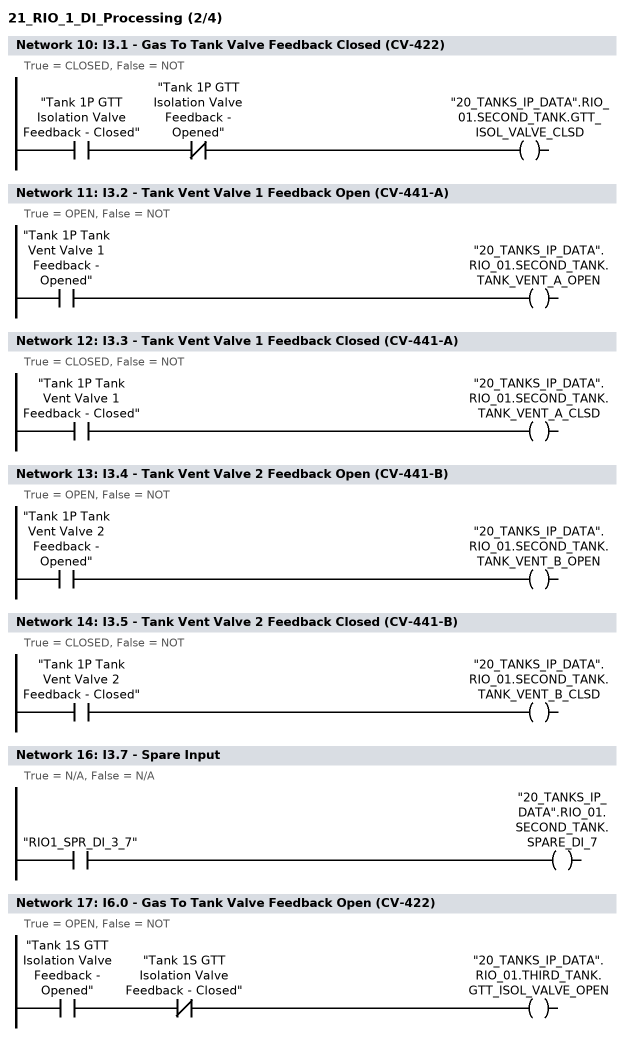
   RUNG wire#powerrail
      Contact( "Tank 1P GTT Isolation Valve Feedback - Closed" )
      I_Contact( "Tank 1P GTT Isolation Valve Feedback - Opened" )
      Coil( "20_TANKS_IP_DATA".RIO_01.SECOND_TANK.GTT_ISOL_VALVE_CLSD )
   END_RUNG
   // the same network as SCL:
   "20_TANKS_IP_DATA".RIO_01.SECOND_TANK.GTT_ISOL_VALVE_CLSD := "Tank 1P GTT Isolation Valve Feedback - Closed" AND NOT "Tank 1P GTT Isolation Valve Feedback - Opened";
END_REGION

REGION Network 11: I3.2 - Tank Vent Valve 1 Feedback Open (CV-441-A)
   // True = OPEN, False = NOT
   RUNG wire#powerrail
      Contact( "Tank 1P Tank Vent Valve 1 Feedback - Opened" )
      Coil( "20_TANKS_IP_DATA".RIO_01.SECOND_TANK.TANK_VENT_A_OPEN )
   END_RUNG
   // the same network as SCL:
   "20_TANKS_IP_DATA".RIO_01.SECOND_TANK.TANK_VENT_A_OPEN := "Tank 1P Tank Vent Valve 1 Feedback - Opened";
END_REGION

REGION Network 12: I3.3 - Tank Vent Valve 1 Feedback Closed (CV-441-A)
   // True = CLOSED, False = NOT
   RUNG wire#powerrail
      Contact( "Tank 1P Tank Vent Valve 1 Feedback - Closed" )
      Coil( "20_TANKS_IP_DATA".RIO_01.SECOND_TANK.TANK_VENT_A_CLSD )
   END_RUNG
   // the same network as SCL:
   "20_TANKS_IP_DATA".RIO_01.SECOND_TANK.TANK_VENT_A_CLSD := "Tank 1P Tank Vent Valve 1 Feedback - Closed";
END_REGION

REGION Network 13: I3.4 - Tank Vent Valve 2 Feedback Open (CV-441-B)
   // True = OPEN, False = NOT
   RUNG wire#powerrail
      Contact( "Tank 1P Tank Vent Valve 2 Feedback - Opened" )
      Coil( "20_TANKS_IP_DATA".RIO_01.SECOND_TANK.TANK_VENT_B_OPEN )
   END_RUNG
   // the same network as SCL:
   "20_TANKS_IP_DATA".RIO_01.SECOND_TANK.TANK_VENT_B_OPEN := "Tank 1P Tank Vent Valve 2 Feedback - Opened";
END_REGION

REGION Network 14: I3.5 - Tank Vent Valve 2 Feedback Closed (CV-441-B)
   // True = CLOSED, False = NOT
   RUNG wire#powerrail
      Contact( "Tank 1P Tank Vent Valve 2 Feedback - Closed" )
      Coil( "20_TANKS_IP_DATA".RIO_01.SECOND_TANK.TANK_VENT_B_CLSD )
   END_RUNG
   // the same network as SCL:
   "20_TANKS_IP_DATA".RIO_01.SECOND_TANK.TANK_VENT_B_CLSD := "Tank 1P Tank Vent Valve 2 Feedback - Closed";
END_REGION

REGION Network 15: I3.6 - Spare Input Accesed from Warning FC
   // True = N/A, False = N/A
END_REGION

REGION Network 16: I3.7 - Spare Input
   // True = N/A, False = N/A
   RUNG wire#powerrail
      Contact( "RIO1_SPR_DI_3_7" )
      Coil( "20_TANKS_IP_DATA".RIO_01.SECOND_TANK.SPARE_DI_7 )
   END_RUNG
   // the same network as SCL:
   "20_TANKS_IP_DATA".RIO_01.SECOND_TANK.SPARE_DI_7 := "RIO1_SPR_DI_3_7";
END_REGION

REGION Network 17: I6.0 - Gas To Tank Valve Feedback Open (CV-422)
   // True = OPEN, False = NOT
   RUNG wire#powerrail
      Contact( "Tank 1S GTT Isolation Valve Feedback - Opened" )
      I_Contact( "Tank 1S GTT Isolation Valve Feedback - Closed" )
      Coil( "20_TANKS_IP_DATA".RIO_01.THIRD_TANK.GTT_ISOL_VALVE_OPEN )
   END_RUNG
   // the same network as SCL:
   "20_TANKS_IP_DATA".RIO_01.THIRD_TANK.GTT_ISOL_VALVE_OPEN := "Tank 1S GTT Isolation Valve Feedback - Opened" AND NOT "Tank 1S GTT Isolation Valve Feedback - Closed";
END_REGION

REGION Network 18: I6.1 - Gas To Tank Valve Feedback Closed (CV-422)
   // True = CLOSED, False = NOT
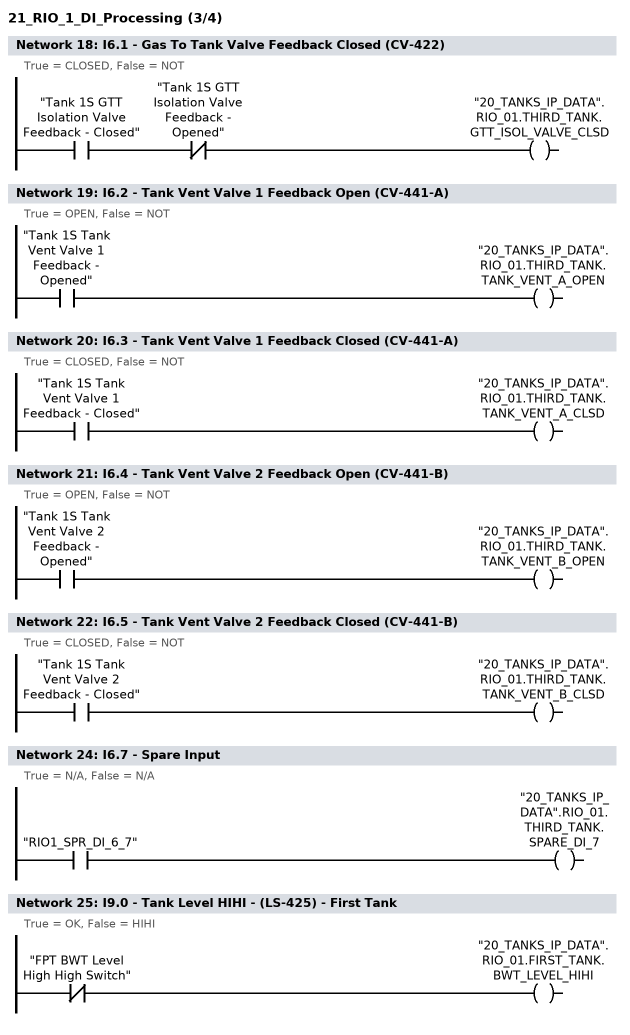
   RUNG wire#powerrail
      Contact( "Tank 1S GTT Isolation Valve Feedback - Closed" )
      I_Contact( "Tank 1S GTT Isolation Valve Feedback - Opened" )
      Coil( "20_TANKS_IP_DATA".RIO_01.THIRD_TANK.GTT_ISOL_VALVE_CLSD )
   END_RUNG
   // the same network as SCL:
   "20_TANKS_IP_DATA".RIO_01.THIRD_TANK.GTT_ISOL_VALVE_CLSD := "Tank 1S GTT Isolation Valve Feedback - Closed" AND NOT "Tank 1S GTT Isolation Valve Feedback - Opened";
END_REGION

REGION Network 19: I6.2 - Tank Vent Valve 1 Feedback Open (CV-441-A)
   // True = OPEN, False = NOT
   RUNG wire#powerrail
      Contact( "Tank 1S Tank Vent Valve 1 Feedback - Opened" )
      Coil( "20_TANKS_IP_DATA".RIO_01.THIRD_TANK.TANK_VENT_A_OPEN )
   END_RUNG
   // the same network as SCL:
   "20_TANKS_IP_DATA".RIO_01.THIRD_TANK.TANK_VENT_A_OPEN := "Tank 1S Tank Vent Valve 1 Feedback - Opened";
END_REGION

REGION Network 20: I6.3 - Tank Vent Valve 1 Feedback Closed (CV-441-A)
   // True = CLOSED, False = NOT
   RUNG wire#powerrail
      Contact( "Tank 1S Tank Vent Valve 1 Feedback - Closed" )
      Coil( "20_TANKS_IP_DATA".RIO_01.THIRD_TANK.TANK_VENT_A_CLSD )
   END_RUNG
   // the same network as SCL:
   "20_TANKS_IP_DATA".RIO_01.THIRD_TANK.TANK_VENT_A_CLSD := "Tank 1S Tank Vent Valve 1 Feedback - Closed";
END_REGION

REGION Network 21: I6.4 - Tank Vent Valve 2 Feedback Open (CV-441-B)
   // True = OPEN, False = NOT
   RUNG wire#powerrail
      Contact( "Tank 1S Tank Vent Valve 2 Feedback - Opened" )
      Coil( "20_TANKS_IP_DATA".RIO_01.THIRD_TANK.TANK_VENT_B_OPEN )
   END_RUNG
   // the same network as SCL:
   "20_TANKS_IP_DATA".RIO_01.THIRD_TANK.TANK_VENT_B_OPEN := "Tank 1S Tank Vent Valve 2 Feedback - Opened";
END_REGION

REGION Network 22: I6.5 - Tank Vent Valve 2 Feedback Closed (CV-441-B)
   // True = CLOSED, False = NOT
   RUNG wire#powerrail
      Contact( "Tank 1S Tank Vent Valve 2 Feedback - Closed" )
      Coil( "20_TANKS_IP_DATA".RIO_01.THIRD_TANK.TANK_VENT_B_CLSD )
   END_RUNG
   // the same network as SCL:
   "20_TANKS_IP_DATA".RIO_01.THIRD_TANK.TANK_VENT_B_CLSD := "Tank 1S Tank Vent Valve 2 Feedback - Closed";
END_REGION

REGION Network 23: I6.6 - Spare Input Accesed from Warning FC
   // True = N/A, False = N/A
END_REGION

REGION Network 24: I6.7 - Spare Input
   // True = N/A, False = N/A
   RUNG wire#powerrail
      Contact( "RIO1_SPR_DI_6_7" )
      Coil( "20_TANKS_IP_DATA".RIO_01.THIRD_TANK.SPARE_DI_7 )
   END_RUNG
   // the same network as SCL:
   "20_TANKS_IP_DATA".RIO_01.THIRD_TANK.SPARE_DI_7 := "RIO1_SPR_DI_6_7";
END_REGION

REGION Network 25: I9.0 - Tank Level HIHI - (LS-425) - First Tank
   // True = OK, False = HIHI
   RUNG wire#powerrail
      I_Contact( "FPT BWT Level High High Switch" )
      Coil( "20_TANKS_IP_DATA".RIO_01.FIRST_TANK.BWT_LEVEL_HIHI )
   END_RUNG
   // the same network as SCL:
   "20_TANKS_IP_DATA".RIO_01.FIRST_TANK.BWT_LEVEL_HIHI := NOT "FPT BWT Level High High Switch";
END_REGION

REGION Network 26: I9.1 - Tank Group Pressure HIHI (PS-436)
   // True = OK, False = HIHI
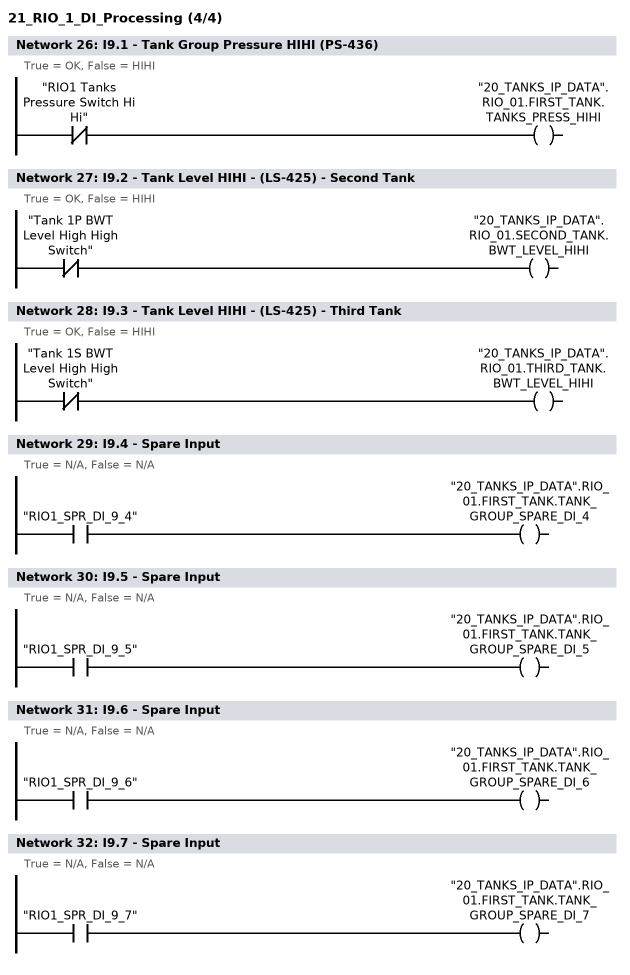
   RUNG wire#powerrail
      I_Contact( "RIO1 Tanks Pressure Switch Hi Hi" )
      Coil( "20_TANKS_IP_DATA".RIO_01.FIRST_TANK.TANKS_PRESS_HIHI )
   END_RUNG
   // the same network as SCL:
   "20_TANKS_IP_DATA".RIO_01.FIRST_TANK.TANKS_PRESS_HIHI := NOT "RIO1 Tanks Pressure Switch Hi Hi";
END_REGION

REGION Network 27: I9.2 - Tank Level HIHI - (LS-425) - Second Tank
   // True = OK, False = HIHI
   RUNG wire#powerrail
      I_Contact( "Tank 1P BWT Level High High Switch" )
      Coil( "20_TANKS_IP_DATA".RIO_01.SECOND_TANK.BWT_LEVEL_HIHI )
   END_RUNG
   // the same network as SCL:
   "20_TANKS_IP_DATA".RIO_01.SECOND_TANK.BWT_LEVEL_HIHI := NOT "Tank 1P BWT Level High High Switch";
END_REGION

REGION Network 28: I9.3 - Tank Level HIHI - (LS-425) - Third Tank
   // True = OK, False = HIHI
   RUNG wire#powerrail
      I_Contact( "Tank 1S BWT Level High High Switch" )
      Coil( "20_TANKS_IP_DATA".RIO_01.THIRD_TANK.BWT_LEVEL_HIHI )
   END_RUNG
   // the same network as SCL:
   "20_TANKS_IP_DATA".RIO_01.THIRD_TANK.BWT_LEVEL_HIHI := NOT "Tank 1S BWT Level High High Switch";
END_REGION

REGION Network 29: I9.4 - Spare Input
   // True = N/A, False = N/A
   RUNG wire#powerrail
      Contact( "RIO1_SPR_DI_9_4" )
      Coil( "20_TANKS_IP_DATA".RIO_01.FIRST_TANK.TANK_GROUP_SPARE_DI_4 )
   END_RUNG
   // the same network as SCL:
   "20_TANKS_IP_DATA".RIO_01.FIRST_TANK.TANK_GROUP_SPARE_DI_4 := "RIO1_SPR_DI_9_4";
END_REGION

REGION Network 30: I9.5 - Spare Input
   // True = N/A, False = N/A
   RUNG wire#powerrail
      Contact( "RIO1_SPR_DI_9_5" )
      Coil( "20_TANKS_IP_DATA".RIO_01.FIRST_TANK.TANK_GROUP_SPARE_DI_5 )
   END_RUNG
   // the same network as SCL:
   "20_TANKS_IP_DATA".RIO_01.FIRST_TANK.TANK_GROUP_SPARE_DI_5 := "RIO1_SPR_DI_9_5";
END_REGION

REGION Network 31: I9.6 - Spare Input
   // True = N/A, False = N/A
   RUNG wire#powerrail
      Contact( "RIO1_SPR_DI_9_6" )
      Coil( "20_TANKS_IP_DATA".RIO_01.FIRST_TANK.TANK_GROUP_SPARE_DI_6 )
   END_RUNG
   // the same network as SCL:
   "20_TANKS_IP_DATA".RIO_01.FIRST_TANK.TANK_GROUP_SPARE_DI_6 := "RIO1_SPR_DI_9_6";
END_REGION

REGION Network 32: I9.7 - Spare Input
   // True = N/A, False = N/A
   RUNG wire#powerrail
      Contact( "RIO1_SPR_DI_9_7" )
      Coil( "20_TANKS_IP_DATA".RIO_01.FIRST_TANK.TANK_GROUP_SPARE_DI_7 )
   END_RUNG
   // the same network as SCL:
   "20_TANKS_IP_DATA".RIO_01.FIRST_TANK.TANK_GROUP_SPARE_DI_7 := "RIO1_SPR_DI_9_7";
END_REGION
END_FUNCTION

FUNCTION "22_RIO_2_DI_Processing" : Void   // FC22, LAD
TITLE = RIO Rack Digital Input Processing (Tank 1 = 2P, Tank 2 = 2S)
{ S7_Optimized_Access := 'TRUE' }
AUTHOR : JRS
VERSION : 0.1
// To process raw inputs prior to code use
BEGIN

REGION Network 1: I15.0 - Gas To Tank Valve Feedback Open (CV-422)
   // True = OPEN, False = NOT
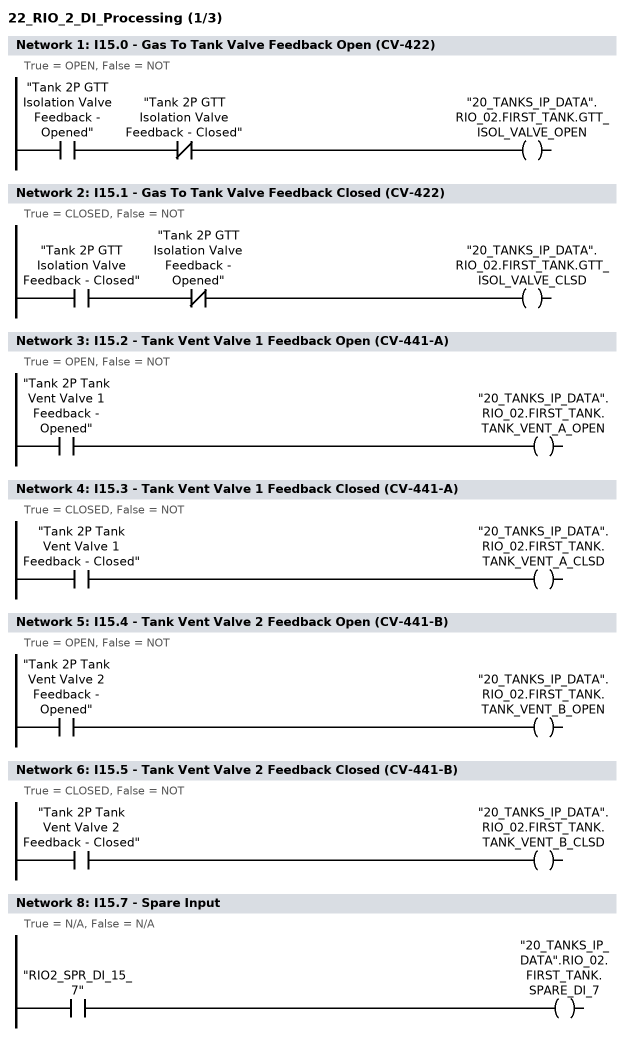
   RUNG wire#powerrail
      Contact( "Tank 2P GTT Isolation Valve Feedback - Opened" )
      I_Contact( "Tank 2P GTT Isolation Valve Feedback - Closed" )
      Coil( "20_TANKS_IP_DATA".RIO_02.FIRST_TANK.GTT_ISOL_VALVE_OPEN )
   END_RUNG
   // the same network as SCL:
   "20_TANKS_IP_DATA".RIO_02.FIRST_TANK.GTT_ISOL_VALVE_OPEN := "Tank 2P GTT Isolation Valve Feedback - Opened" AND NOT "Tank 2P GTT Isolation Valve Feedback - Closed";
END_REGION

REGION Network 2: I15.1 - Gas To Tank Valve Feedback Closed (CV-422)
   // True = CLOSED, False = NOT
   RUNG wire#powerrail
      Contact( "Tank 2P GTT Isolation Valve Feedback - Closed" )
      I_Contact( "Tank 2P GTT Isolation Valve Feedback - Opened" )
      Coil( "20_TANKS_IP_DATA".RIO_02.FIRST_TANK.GTT_ISOL_VALVE_CLSD )
   END_RUNG
   // the same network as SCL:
   "20_TANKS_IP_DATA".RIO_02.FIRST_TANK.GTT_ISOL_VALVE_CLSD := "Tank 2P GTT Isolation Valve Feedback - Closed" AND NOT "Tank 2P GTT Isolation Valve Feedback - Opened";
END_REGION

REGION Network 3: I15.2 - Tank Vent Valve 1 Feedback Open (CV-441-A)
   // True = OPEN, False = NOT
   RUNG wire#powerrail
      Contact( "Tank 2P Tank Vent Valve 1 Feedback - Opened" )
      Coil( "20_TANKS_IP_DATA".RIO_02.FIRST_TANK.TANK_VENT_A_OPEN )
   END_RUNG
   // the same network as SCL:
   "20_TANKS_IP_DATA".RIO_02.FIRST_TANK.TANK_VENT_A_OPEN := "Tank 2P Tank Vent Valve 1 Feedback - Opened";
END_REGION

REGION Network 4: I15.3 - Tank Vent Valve 1 Feedback Closed (CV-441-A)
   // True = CLOSED, False = NOT
   RUNG wire#powerrail
      Contact( "Tank 2P Tank Vent Valve 1 Feedback - Closed" )
      Coil( "20_TANKS_IP_DATA".RIO_02.FIRST_TANK.TANK_VENT_A_CLSD )
   END_RUNG
   // the same network as SCL:
   "20_TANKS_IP_DATA".RIO_02.FIRST_TANK.TANK_VENT_A_CLSD := "Tank 2P Tank Vent Valve 1 Feedback - Closed";
END_REGION

REGION Network 5: I15.4 - Tank Vent Valve 2 Feedback Open (CV-441-B)
   // True = OPEN, False = NOT
   RUNG wire#powerrail
      Contact( "Tank 2P Tank Vent Valve 2 Feedback - Opened" )
      Coil( "20_TANKS_IP_DATA".RIO_02.FIRST_TANK.TANK_VENT_B_OPEN )
   END_RUNG
   // the same network as SCL:
   "20_TANKS_IP_DATA".RIO_02.FIRST_TANK.TANK_VENT_B_OPEN := "Tank 2P Tank Vent Valve 2 Feedback - Opened";
END_REGION

REGION Network 6: I15.5 - Tank Vent Valve 2 Feedback Closed (CV-441-B)
   // True = CLOSED, False = NOT
   RUNG wire#powerrail
      Contact( "Tank 2P Tank Vent Valve 2 Feedback - Closed" )
      Coil( "20_TANKS_IP_DATA".RIO_02.FIRST_TANK.TANK_VENT_B_CLSD )
   END_RUNG
   // the same network as SCL:
   "20_TANKS_IP_DATA".RIO_02.FIRST_TANK.TANK_VENT_B_CLSD := "Tank 2P Tank Vent Valve 2 Feedback - Closed";
END_REGION

REGION Network 7: I15.6 - Spare Input Accesed from Warning FC
   // True = N/A, False = N/A
END_REGION

REGION Network 8: I15.7 - Spare Input
   // True = N/A, False = N/A
   RUNG wire#powerrail
      Contact( "RIO2_SPR_DI_15_7" )
      Coil( "20_TANKS_IP_DATA".RIO_02.FIRST_TANK.SPARE_DI_7 )
   END_RUNG
   // the same network as SCL:
   "20_TANKS_IP_DATA".RIO_02.FIRST_TANK.SPARE_DI_7 := "RIO2_SPR_DI_15_7";
END_REGION

REGION Network 9: I18.0 - Gas To Tank Valve Feedback Open (CV-422)
   // True = OPEN, False = NOT
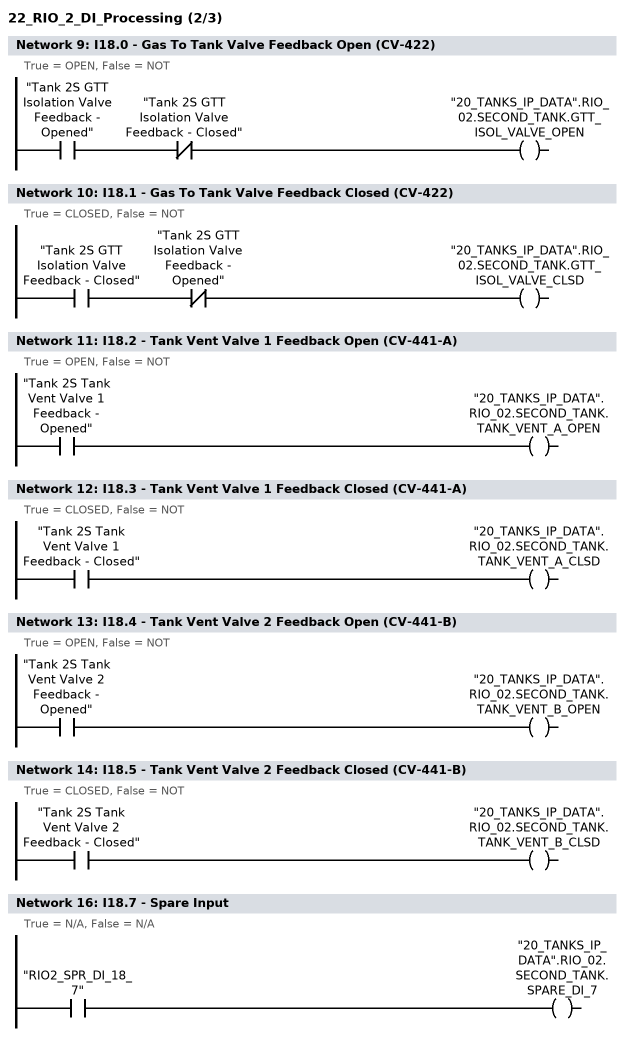
   RUNG wire#powerrail
      Contact( "Tank 2S GTT Isolation Valve Feedback - Opened" )
      I_Contact( "Tank 2S GTT Isolation Valve Feedback - Closed" )
      Coil( "20_TANKS_IP_DATA".RIO_02.SECOND_TANK.GTT_ISOL_VALVE_OPEN )
   END_RUNG
   // the same network as SCL:
   "20_TANKS_IP_DATA".RIO_02.SECOND_TANK.GTT_ISOL_VALVE_OPEN := "Tank 2S GTT Isolation Valve Feedback - Opened" AND NOT "Tank 2S GTT Isolation Valve Feedback - Closed";
END_REGION

REGION Network 10: I18.1 - Gas To Tank Valve Feedback Closed (CV-422)
   // True = CLOSED, False = NOT
   RUNG wire#powerrail
      Contact( "Tank 2S GTT Isolation Valve Feedback - Closed" )
      I_Contact( "Tank 2S GTT Isolation Valve Feedback - Opened" )
      Coil( "20_TANKS_IP_DATA".RIO_02.SECOND_TANK.GTT_ISOL_VALVE_CLSD )
   END_RUNG
   // the same network as SCL:
   "20_TANKS_IP_DATA".RIO_02.SECOND_TANK.GTT_ISOL_VALVE_CLSD := "Tank 2S GTT Isolation Valve Feedback - Closed" AND NOT "Tank 2S GTT Isolation Valve Feedback - Opened";
END_REGION

REGION Network 11: I18.2 - Tank Vent Valve 1 Feedback Open (CV-441-A)
   // True = OPEN, False = NOT
   RUNG wire#powerrail
      Contact( "Tank 2S Tank Vent Valve 1 Feedback - Opened" )
      Coil( "20_TANKS_IP_DATA".RIO_02.SECOND_TANK.TANK_VENT_A_OPEN )
   END_RUNG
   // the same network as SCL:
   "20_TANKS_IP_DATA".RIO_02.SECOND_TANK.TANK_VENT_A_OPEN := "Tank 2S Tank Vent Valve 1 Feedback - Opened";
END_REGION

REGION Network 12: I18.3 - Tank Vent Valve 1 Feedback Closed (CV-441-A)
   // True = CLOSED, False = NOT
   RUNG wire#powerrail
      Contact( "Tank 2S Tank Vent Valve 1 Feedback - Closed" )
      Coil( "20_TANKS_IP_DATA".RIO_02.SECOND_TANK.TANK_VENT_A_CLSD )
   END_RUNG
   // the same network as SCL:
   "20_TANKS_IP_DATA".RIO_02.SECOND_TANK.TANK_VENT_A_CLSD := "Tank 2S Tank Vent Valve 1 Feedback - Closed";
END_REGION

REGION Network 13: I18.4 - Tank Vent Valve 2 Feedback Open (CV-441-B)
   // True = OPEN, False = NOT
   RUNG wire#powerrail
      Contact( "Tank 2S Tank Vent Valve 2 Feedback - Opened" )
      Coil( "20_TANKS_IP_DATA".RIO_02.SECOND_TANK.TANK_VENT_B_OPEN )
   END_RUNG
   // the same network as SCL:
   "20_TANKS_IP_DATA".RIO_02.SECOND_TANK.TANK_VENT_B_OPEN := "Tank 2S Tank Vent Valve 2 Feedback - Opened";
END_REGION

REGION Network 14: I18.5 - Tank Vent Valve 2 Feedback Closed (CV-441-B)
   // True = CLOSED, False = NOT
   RUNG wire#powerrail
      Contact( "Tank 2S Tank Vent Valve 2 Feedback - Closed" )
      Coil( "20_TANKS_IP_DATA".RIO_02.SECOND_TANK.TANK_VENT_B_CLSD )
   END_RUNG
   // the same network as SCL:
   "20_TANKS_IP_DATA".RIO_02.SECOND_TANK.TANK_VENT_B_CLSD := "Tank 2S Tank Vent Valve 2 Feedback - Closed";
END_REGION

REGION Network 15: I18.6 - Spare Input Accesed from Warning FC
   // True = N/A, False = N/A
END_REGION

REGION Network 16: I18.7 - Spare Input
   // True = N/A, False = N/A
   RUNG wire#powerrail
      Contact( "RIO2_SPR_DI_18_7" )
      Coil( "20_TANKS_IP_DATA".RIO_02.SECOND_TANK.SPARE_DI_7 )
   END_RUNG
   // the same network as SCL:
   "20_TANKS_IP_DATA".RIO_02.SECOND_TANK.SPARE_DI_7 := "RIO2_SPR_DI_18_7";
END_REGION

REGION Network 17: I21.0 - Tank Level HIHI - (LS-425) - First Tank
   // True = OK, False = HIHI
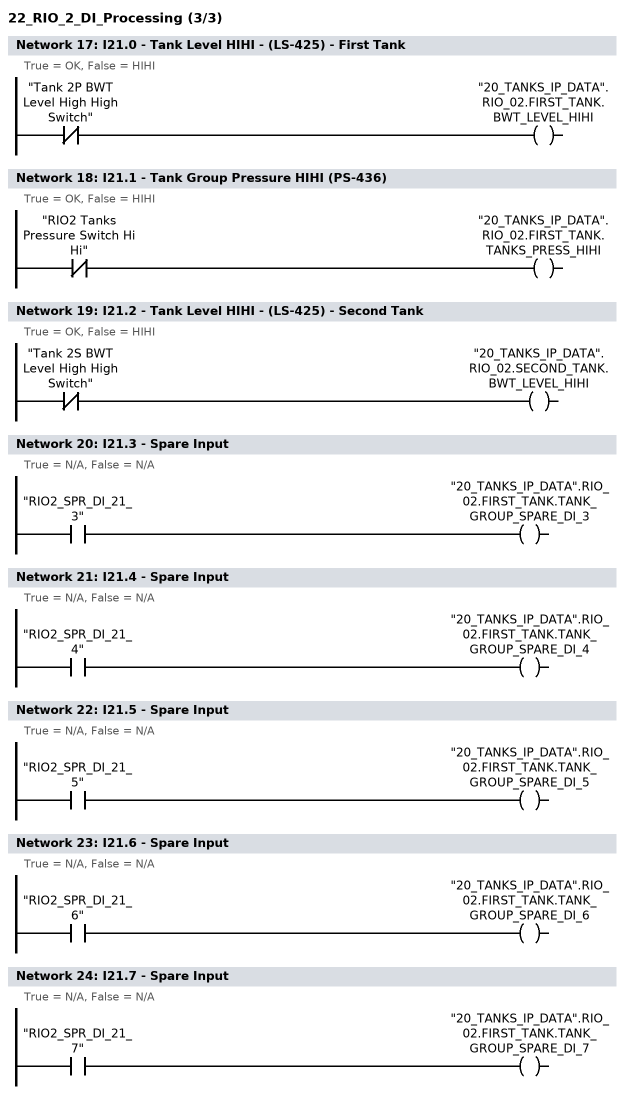
   RUNG wire#powerrail
      I_Contact( "Tank 2P BWT Level High High Switch" )
      Coil( "20_TANKS_IP_DATA".RIO_02.FIRST_TANK.BWT_LEVEL_HIHI )
   END_RUNG
   // the same network as SCL:
   "20_TANKS_IP_DATA".RIO_02.FIRST_TANK.BWT_LEVEL_HIHI := NOT "Tank 2P BWT Level High High Switch";
END_REGION
